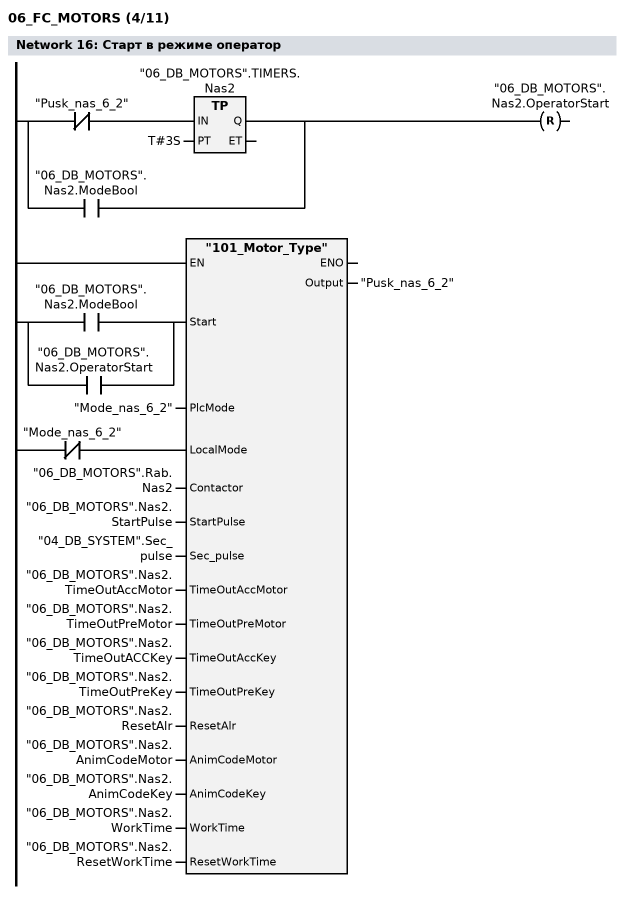
   "06_DB_MOTORS".TIMERS.Nas2.TP(IN := NOT "Pusk_nas_6_2", PT := T#3S);
   IF "06_DB_MOTORS".TIMERS.Nas2.Q OR "06_DB_MOTORS".Nas2.ModeBool THEN
       "06_DB_MOTORS".Nas2.OperatorStart := FALSE;
   END_IF;
   "101_Motor_Type"(Start := "06_DB_MOTORS".Nas2.ModeBool OR "06_DB_MOTORS".Nas2.OperatorStart,
                    PlcMode := "Mode_nas_6_2",
                    LocalMode := NOT "Mode_nas_6_2",
                    Contactor := "06_DB_MOTORS".Rab.Nas2,
                    StartPulse := "06_DB_MOTORS".Nas2.StartPulse,
                    Sec_pulse := "04_DB_SYSTEM".Sec_pulse,
                    TimeOutAccMotor := "06_DB_MOTORS".Nas2.TimeOutAccMotor,
                    TimeOutPreMotor := "06_DB_MOTORS".Nas2.TimeOutPreMotor,
                    TimeOutAccKey := "06_DB_MOTORS".Nas2.TimeOutACCKey,
                    TimeOutPreKey := "06_DB_MOTORS".Nas2.TimeOutPreKey,
                    ResetAlr := "06_DB_MOTORS".Nas2.ResetAlr,
                    AnimCodeMotor := "06_DB_MOTORS".Nas2.AnimCodeMotor,
                    AnimCodeKey := "06_DB_MOTORS".Nas2.AnimCodeKey,
                    WorkTime := "06_DB_MOTORS".Nas2.WorkTime,
                    ResetWorkTime := "06_DB_MOTORS".Nas2.ResetWorkTime,
                    Output => "Pusk_nas_6_2");
END_REGION

REGION Network 17: Старт в режиме оператор
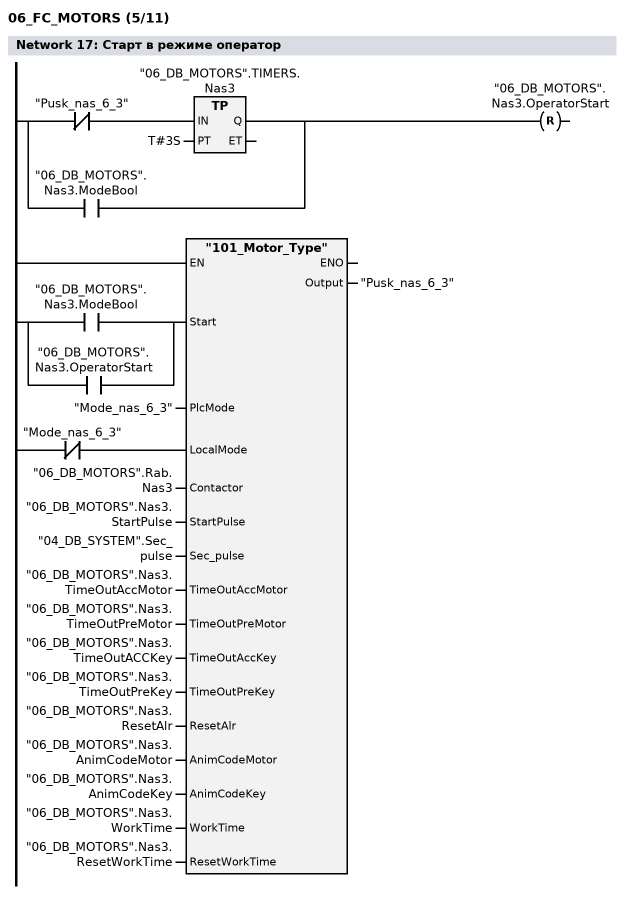
   "06_DB_MOTORS".TIMERS.Nas3.TP(IN := NOT "Pusk_nas_6_3", PT := T#3S);
   IF "06_DB_MOTORS".TIMERS.Nas3.Q OR "06_DB_MOTORS".Nas3.ModeBool THEN
       "06_DB_MOTORS".Nas3.OperatorStart := FALSE;
   END_IF;
   "101_Motor_Type"(Start := "06_DB_MOTORS".Nas3.ModeBool OR "06_DB_MOTORS".Nas3.OperatorStart,
                    PlcMode := "Mode_nas_6_3",
                    LocalMode := NOT "Mode_nas_6_3",
                    Contactor := "06_DB_MOTORS".Rab.Nas3,
                    StartPulse := "06_DB_MOTORS".Nas3.StartPulse,
                    Sec_pulse := "04_DB_SYSTEM".Sec_pulse,
                    TimeOutAccMotor := "06_DB_MOTORS".Nas3.TimeOutAccMotor,
                    TimeOutPreMotor := "06_DB_MOTORS".Nas3.TimeOutPreMotor,
                    TimeOutAccKey := "06_DB_MOTORS".Nas3.TimeOutACCKey,
                    TimeOutPreKey := "06_DB_MOTORS".Nas3.TimeOutPreKey,
                    ResetAlr := "06_DB_MOTORS".Nas3.ResetAlr,
                    AnimCodeMotor := "06_DB_MOTORS".Nas3.AnimCodeMotor,
                    AnimCodeKey := "06_DB_MOTORS".Nas3.AnimCodeKey,
                    WorkTime := "06_DB_MOTORS".Nas3.WorkTime,
                    ResetWorkTime := "06_DB_MOTORS".Nas3.ResetWorkTime,
                    Output => "Pusk_nas_6_3");
END_REGION

REGION Network 18: Старт в режиме оператор
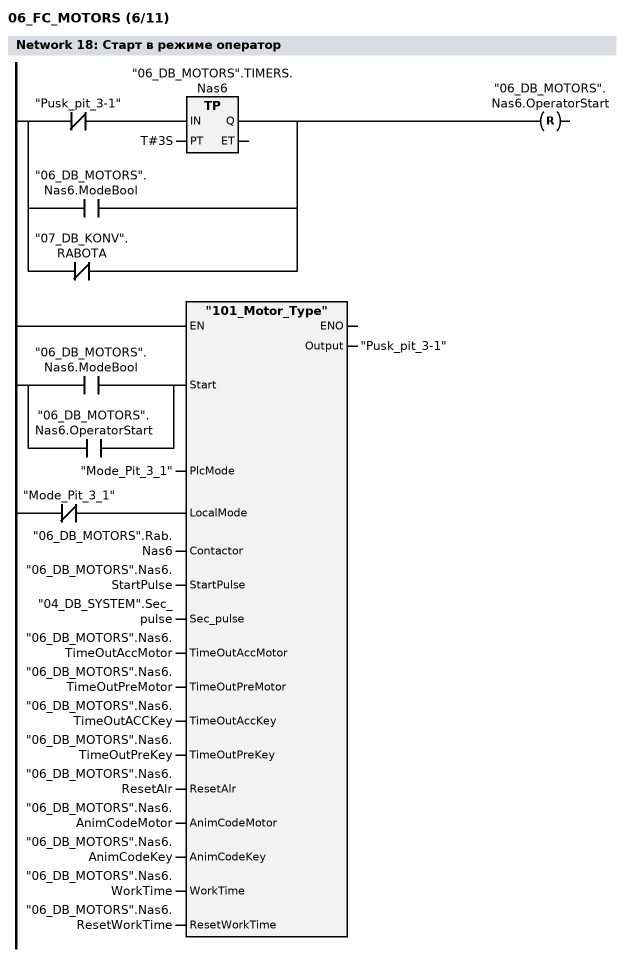
   "06_DB_MOTORS".TIMERS.Nas6.TP(IN := NOT "Pusk_pit_3-1", PT := T#3S);
   IF "06_DB_MOTORS".TIMERS.Nas6.Q OR "06_DB_MOTORS".Nas6.ModeBool OR NOT "07_DB_KONV".RABOTA THEN
       "06_DB_MOTORS".Nas6.OperatorStart := FALSE;
   END_IF;
   "101_Motor_Type"(Start := "06_DB_MOTORS".Nas6.ModeBool OR "06_DB_MOTORS".Nas6.OperatorStart,
                    PlcMode := "Mode_Pit_3_1",
                    LocalMode := NOT "Mode_Pit_3_1",
                    Contactor := "06_DB_MOTORS".Rab.Nas6,
                    StartPulse := "06_DB_MOTORS".Nas6.StartPulse,
                    Sec_pulse := "04_DB_SYSTEM".Sec_pulse,
                    TimeOutAccMotor := "06_DB_MOTORS".Nas6.TimeOutAccMotor,
                    TimeOutPreMotor := "06_DB_MOTORS".Nas6.TimeOutPreMotor,
                    TimeOutAccKey := "06_DB_MOTORS".Nas6.TimeOutACCKey,
                    TimeOutPreKey := "06_DB_MOTORS".Nas6.TimeOutPreKey,
                    ResetAlr := "06_DB_MOTORS".Nas6.ResetAlr,
                    AnimCodeMotor := "06_DB_MOTORS".Nas6.AnimCodeMotor,
                    AnimCodeKey := "06_DB_MOTORS".Nas6.AnimCodeKey,
                    WorkTime := "06_DB_MOTORS".Nas6.WorkTime,
                    ResetWorkTime := "06_DB_MOTORS".Nas6.ResetWorkTime,
                    Output => "Pusk_pit_3-1");
END_REGION

REGION Network 19: Старт в режиме оператор
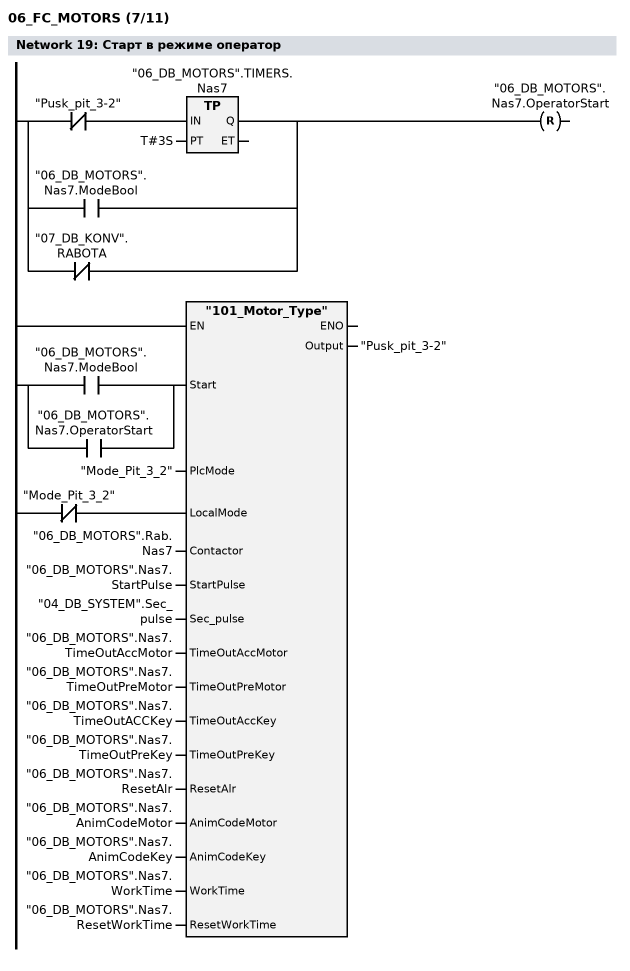
   "06_DB_MOTORS".TIMERS.Nas7.TP(IN := NOT "Pusk_pit_3-2", PT := T#3S);
   IF "06_DB_MOTORS".TIMERS.Nas7.Q OR "06_DB_MOTORS".Nas7.ModeBool OR NOT "07_DB_KONV".RABOTA THEN
       "06_DB_MOTORS".Nas7.OperatorStart := FALSE;
   END_IF;
   "101_Motor_Type"(Start := "06_DB_MOTORS".Nas7.ModeBool OR "06_DB_MOTORS".Nas7.OperatorStart,
                    PlcMode := "Mode_Pit_3_2",
                    LocalMode := NOT "Mode_Pit_3_2",
                    Contactor := "06_DB_MOTORS".Rab.Nas7,
                    StartPulse := "06_DB_MOTORS".Nas7.StartPulse,
                    Sec_pulse := "04_DB_SYSTEM".Sec_pulse,
                    TimeOutAccMotor := "06_DB_MOTORS".Nas7.TimeOutAccMotor,
                    TimeOutPreMotor := "06_DB_MOTORS".Nas7.TimeOutPreMotor,
                    TimeOutAccKey := "06_DB_MOTORS".Nas7.TimeOutACCKey,
                    TimeOutPreKey := "06_DB_MOTORS".Nas7.TimeOutPreKey,
                    ResetAlr := "06_DB_MOTORS".Nas7.ResetAlr,
                    AnimCodeMotor := "06_DB_MOTORS".Nas7.AnimCodeMotor,
                    AnimCodeKey := "06_DB_MOTORS".Nas7.AnimCodeKey,
                    WorkTime := "06_DB_MOTORS".Nas7.WorkTime,
                    ResetWorkTime := "06_DB_MOTORS".Nas7.ResetWorkTime,
                    Output => "Pusk_pit_3-2");
END_REGION

REGION Network 20: Старт в режиме оператор
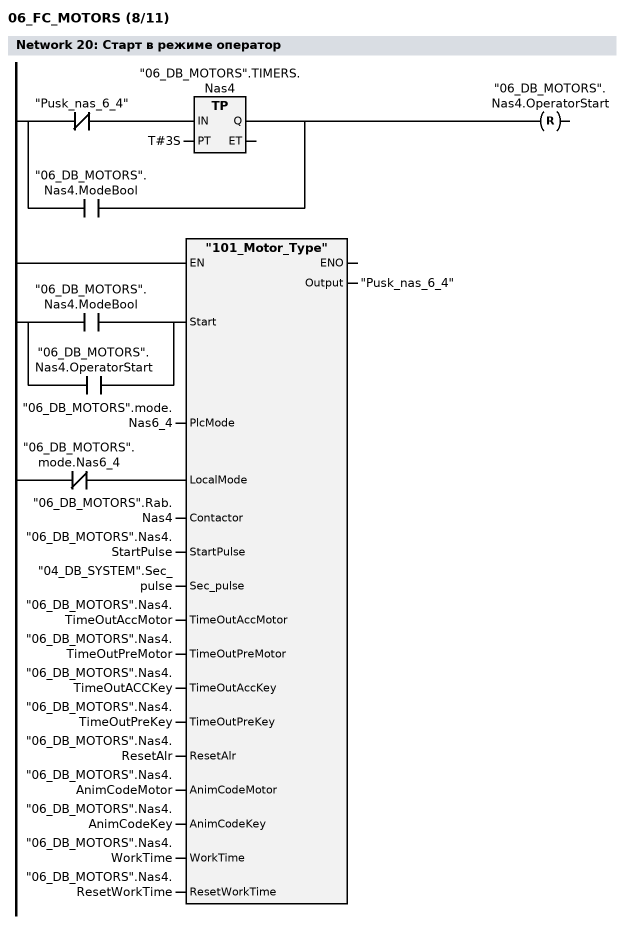
   "06_DB_MOTORS".TIMERS.Nas4.TP(IN := NOT "Pusk_nas_6_4", PT := T#3S);
   IF "06_DB_MOTORS".TIMERS.Nas4.Q OR "06_DB_MOTORS".Nas4.ModeBool THEN
       "06_DB_MOTORS".Nas4.OperatorStart := FALSE;
   END_IF;
   "101_Motor_Type"(Start := "06_DB_MOTORS".Nas4.ModeBool OR "06_DB_MOTORS".Nas4.OperatorStart,
                    PlcMode := "06_DB_MOTORS".mode.Nas6_4,
                    LocalMode := NOT "06_DB_MOTORS".mode.Nas6_4,
                    Contactor := "06_DB_MOTORS".Rab.Nas4,
                    StartPulse := "06_DB_MOTORS".Nas4.StartPulse,
                    Sec_pulse := "04_DB_SYSTEM".Sec_pulse,
                    TimeOutAccMotor := "06_DB_MOTORS".Nas4.TimeOutAccMotor,
                    TimeOutPreMotor := "06_DB_MOTORS".Nas4.TimeOutPreMotor,
                    TimeOutAccKey := "06_DB_MOTORS".Nas4.TimeOutACCKey,
                    TimeOutPreKey := "06_DB_MOTORS".Nas4.TimeOutPreKey,
                    ResetAlr := "06_DB_MOTORS".Nas4.ResetAlr,
                    AnimCodeMotor := "06_DB_MOTORS".Nas4.AnimCodeMotor,
                    AnimCodeKey := "06_DB_MOTORS".Nas4.AnimCodeKey,
                    WorkTime := "06_DB_MOTORS".Nas4.WorkTime,
                    ResetWorkTime := "06_DB_MOTORS".Nas4.ResetWorkTime,
                    Output => "Pusk_nas_6_4");
END_REGION

REGION Network 21: Старт в режиме оператор
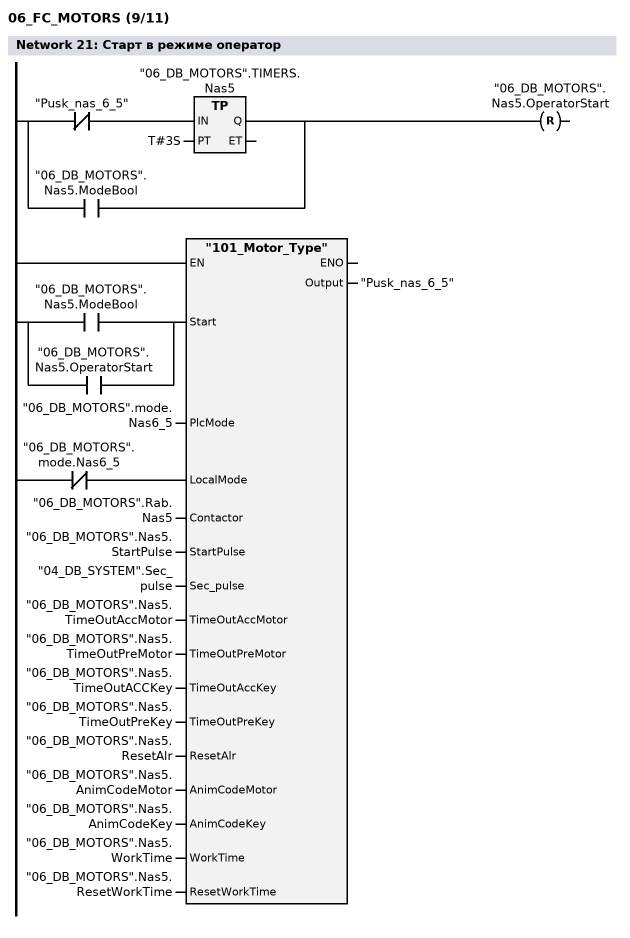
   "06_DB_MOTORS".TIMERS.Nas5.TP(IN := NOT "Pusk_nas_6_5", PT := T#3S);
   IF "06_DB_MOTORS".TIMERS.Nas5.Q OR "06_DB_MOTORS".Nas5.ModeBool THEN
       "06_DB_MOTORS".Nas5.OperatorStart := FALSE;
   END_IF;
   "101_Motor_Type"(Start := "06_DB_MOTORS".Nas5.ModeBool OR "06_DB_MOTORS".Nas5.OperatorStart,
                    PlcMode := "06_DB_MOTORS".mode.Nas6_5,
                    LocalMode := NOT "06_DB_MOTORS".mode.Nas6_5,
                    Contactor := "06_DB_MOTORS".Rab.Nas5,
                    StartPulse := "06_DB_MOTORS".Nas5.StartPulse,
                    Sec_pulse := "04_DB_SYSTEM".Sec_pulse,
                    TimeOutAccMotor := "06_DB_MOTORS".Nas5.TimeOutAccMotor,
                    TimeOutPreMotor := "06_DB_MOTORS".Nas5.TimeOutPreMotor,
                    TimeOutAccKey := "06_DB_MOTORS".Nas5.TimeOutACCKey,
                    TimeOutPreKey := "06_DB_MOTORS".Nas5.TimeOutPreKey,
                    ResetAlr := "06_DB_MOTORS".Nas5.ResetAlr,
                    AnimCodeMotor := "06_DB_MOTORS".Nas5.AnimCodeMotor,
                    AnimCodeKey := "06_DB_MOTORS".Nas5.AnimCodeKey,
                    WorkTime := "06_DB_MOTORS".Nas5.WorkTime,
                    ResetWorkTime := "06_DB_MOTORS".Nas5.ResetWorkTime,
                    Output => "Pusk_nas_6_5");
END_REGION

REGION Network 23: Старт в режиме оператор
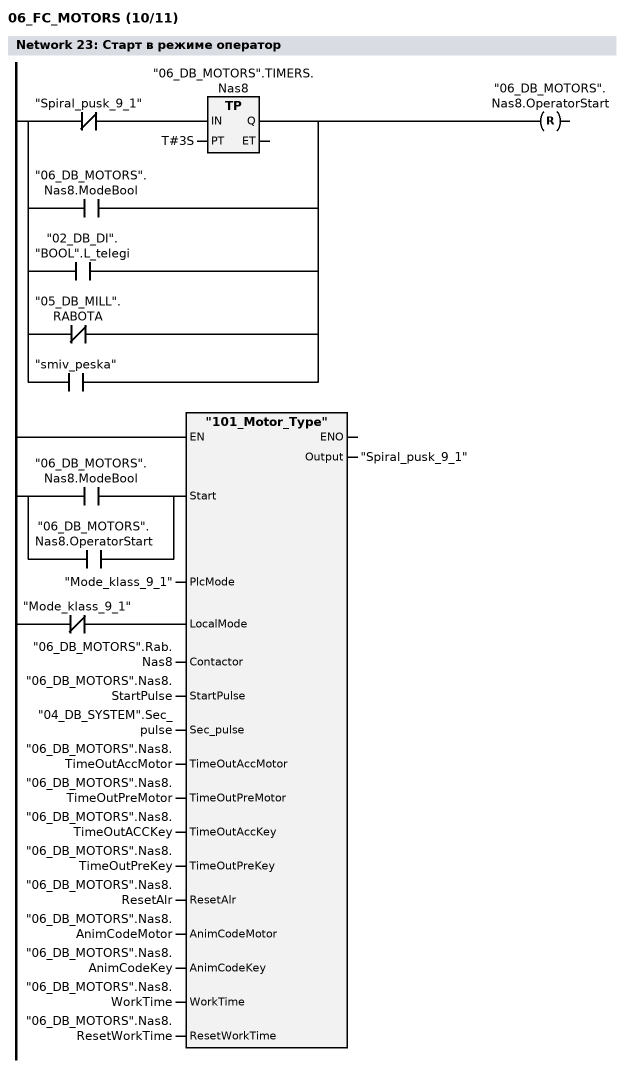
   "06_DB_MOTORS".TIMERS.Nas8.TP(IN := NOT "Spiral_pusk_9_1", PT := T#3S);
   IF "06_DB_MOTORS".TIMERS.Nas8.Q OR "06_DB_MOTORS".Nas8.ModeBool OR "02_DB_DI"."BOOL".L_telegi OR NOT "05_DB_MILL".RABOTA OR "smiv_peska" THEN
       "06_DB_MOTORS".Nas8.OperatorStart := FALSE;
   END_IF;
   "101_Motor_Type"(Start := "06_DB_MOTORS".Nas8.ModeBool OR "06_DB_MOTORS".Nas8.OperatorStart,
                    PlcMode := "Mode_klass_9_1",
                    LocalMode := NOT "Mode_klass_9_1",
                    Contactor := "06_DB_MOTORS".Rab.Nas8,
                    StartPulse := "06_DB_MOTORS".Nas8.StartPulse,
                    Sec_pulse := "04_DB_SYSTEM".Sec_pulse,
                    TimeOutAccMotor := "06_DB_MOTORS".Nas8.TimeOutAccMotor,
                    TimeOutPreMotor := "06_DB_MOTORS".Nas8.TimeOutPreMotor,
                    TimeOutAccKey := "06_DB_MOTORS".Nas8.TimeOutACCKey,
                    TimeOutPreKey := "06_DB_MOTORS".Nas8.TimeOutPreKey,
                    ResetAlr := "06_DB_MOTORS".Nas8.ResetAlr,
                    AnimCodeMotor := "06_DB_MOTORS".Nas8.AnimCodeMotor,
                    AnimCodeKey := "06_DB_MOTORS".Nas8.AnimCodeKey,
                    WorkTime := "06_DB_MOTORS".Nas8.WorkTime,
                    ResetWorkTime := "06_DB_MOTORS".Nas8.ResetWorkTime,
                    Output => "Spiral_pusk_9_1");
END_REGION

REGION Network 24: Старт в режиме оператор
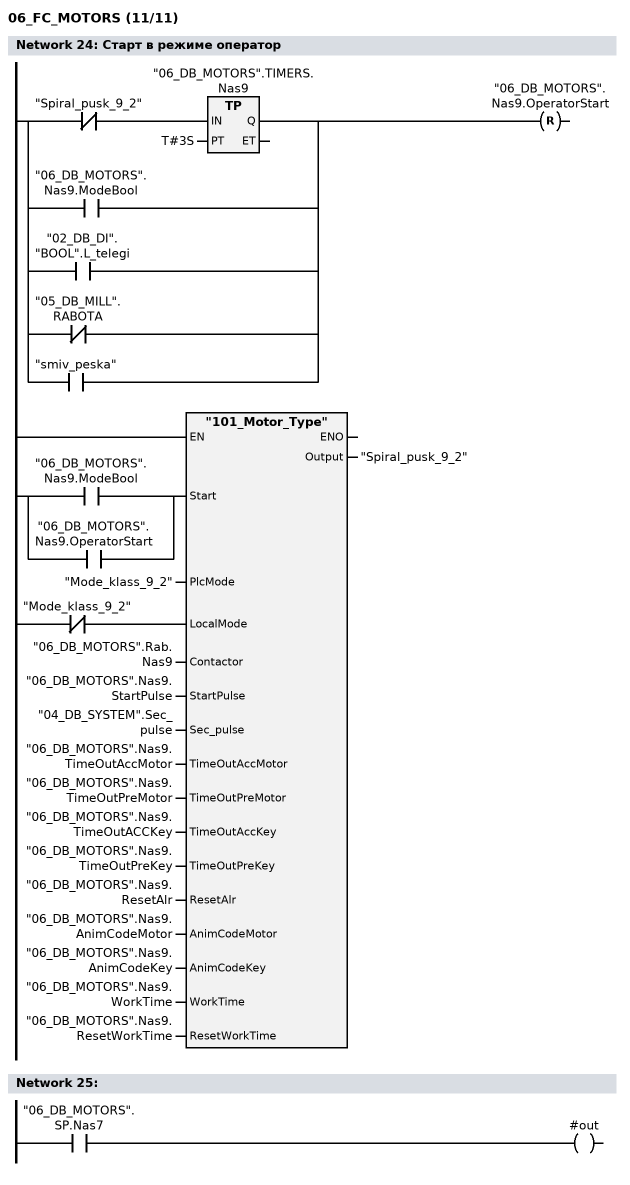
   "06_DB_MOTORS".TIMERS.Nas9.TP(IN := NOT "Spiral_pusk_9_2", PT := T#3S);
   IF "06_DB_MOTORS".TIMERS.Nas9.Q OR "06_DB_MOTORS".Nas9.ModeBool OR "02_DB_DI"."BOOL".L_telegi OR NOT "05_DB_MILL".RABOTA OR "smiv_peska" THEN
       "06_DB_MOTORS".Nas9.OperatorStart := FALSE;
   END_IF;
   "101_Motor_Type"(Start := "06_DB_MOTORS".Nas9.ModeBool OR "06_DB_MOTORS".Nas9.OperatorStart,
                    PlcMode := "Mode_klass_9_2",
                    LocalMode := NOT "Mode_klass_9_2",
                    Contactor := "06_DB_MOTORS".Rab.Nas9,
                    StartPulse := "06_DB_MOTORS".Nas9.StartPulse,
                    Sec_pulse := "04_DB_SYSTEM".Sec_pulse,
                    TimeOutAccMotor := "06_DB_MOTORS".Nas9.TimeOutAccMotor,
                    TimeOutPreMotor := "06_DB_MOTORS".Nas9.TimeOutPreMotor,
                    TimeOutAccKey := "06_DB_MOTORS".Nas9.TimeOutACCKey,
                    TimeOutPreKey := "06_DB_MOTORS".Nas9.TimeOutPreKey,
                    ResetAlr := "06_DB_MOTORS".Nas9.ResetAlr,
                    AnimCodeMotor := "06_DB_MOTORS".Nas9.AnimCodeMotor,
                    AnimCodeKey := "06_DB_MOTORS".Nas9.AnimCodeKey,
                    WorkTime := "06_DB_MOTORS".Nas9.WorkTime,
                    ResetWorkTime := "06_DB_MOTORS".Nas9.ResetWorkTime,
                    Output => "Spiral_pusk_9_2");
END_REGION

REGION Network 25
   RUNG wire#powerrail
      Contact( "06_DB_MOTORS".SP.Nas7 )
      Coil( #out )
   END_RUNG
   // the same network as SCL:
   #out := "06_DB_MOTORS".SP.Nas7;
END_REGION
END_FUNCTION

FUNCTION "09_alarm" : Void   // FC9, LAD
{ S7_Optimized_Access := 'TRUE' }
VERSION : 0.1
   VAR_TEMP   // added for the SCL form of the ladder/FBD networks
      _w1 : Bool;
      _w2 : Bool;
      _w3 : Bool;
      _w4 : Bool;
      _w5 : Bool;
      _w6 : Bool;
      _w7 : Bool;
      _w8 : Bool;
      _w9 : Bool;
      _w10 : Bool;
      _w11 : Bool;
      _w12 : Bool;
      _w13 : Bool;
      _w14 : Bool;
      _w15 : Bool;
      _w16 : Bool;
   END_VAR
BEGIN

REGION Network 1
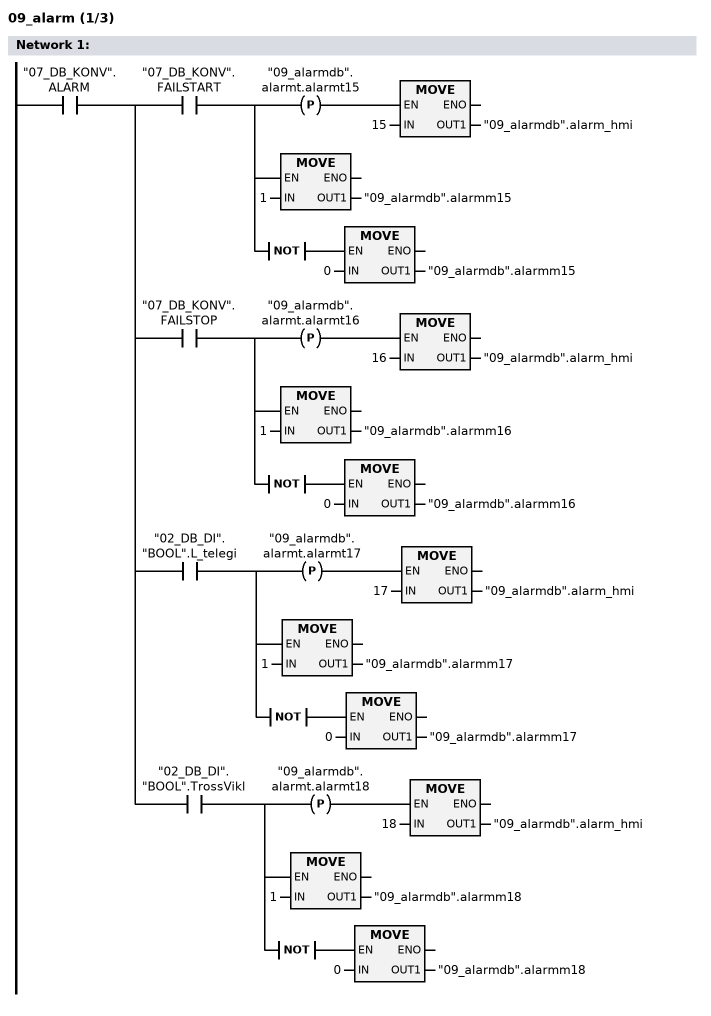
   RUNG wire#powerrail
      Contact( "07_DB_KONV".ALARM )
      wire#w1
      Contact( "07_DB_KONV".FAILSTART )
      wire#w2
      P_Trig( "09_alarmdb".alarmt.alarmt15 )
      Move(in := 15, out1 => "09_alarmdb".alarm_hmi)
   END_RUNG
   RUNG wire#w2
      Move(in := 1, out1 => "09_alarmdb".alarmm15)
   END_RUNG
   RUNG wire#w2
      Not()
      Move(in := 0, out1 => "09_alarmdb".alarmm15)
   END_RUNG
   RUNG wire#w1
      Contact( "07_DB_KONV".FAILSTOP )
      wire#w3
      P_Trig( "09_alarmdb".alarmt.alarmt16 )
      Move(in := 16, out1 => "09_alarmdb".alarm_hmi)
   END_RUNG
   RUNG wire#w3
      Move(in := 1, out1 => "09_alarmdb".alarmm16)
   END_RUNG
   RUNG wire#w3
      Not()
      Move(in := 0, out1 => "09_alarmdb".alarmm16)
   END_RUNG
   RUNG wire#w1
      Contact( "02_DB_DI"."BOOL".L_telegi )
      wire#w4
      P_Trig( "09_alarmdb".alarmt.alarmt17 )
      Move(in := 17, out1 => "09_alarmdb".alarm_hmi)
   END_RUNG
   RUNG wire#w4
      Move(in := 1, out1 => "09_alarmdb".alarmm17)
   END_RUNG
   RUNG wire#w4
      Not()
      Move(in := 0, out1 => "09_alarmdb".alarmm17)
   END_RUNG
   RUNG wire#w1
      Contact( "02_DB_DI"."BOOL".TrossVikl )
      wire#w5
      P_Trig( "09_alarmdb".alarmt.alarmt18 )
      Move(in := 18, out1 => "09_alarmdb".alarm_hmi)
   END_RUNG
   RUNG wire#w5
      Move(in := 1, out1 => "09_alarmdb".alarmm18)
   END_RUNG
   RUNG wire#w5
      Not()
      Move(in := 0, out1 => "09_alarmdb".alarmm18)
   END_RUNG
   // the same network as SCL:
   #_w1 := "07_DB_KONV".ALARM AND "07_DB_KONV".FAILSTART;
   #_w2 := #_w1 AND NOT "09_alarmdb".alarmt.alarmt15;   // rising edge
   "09_alarmdb".alarmt.alarmt15 := #_w1;
   IF #_w2 THEN "09_alarmdb".alarm_hmi := 15; END_IF;
   IF #_w1 THEN "09_alarmdb".alarmm15 := 1; END_IF;
   IF NOT #_w1 THEN "09_alarmdb".alarmm15 := 0; END_IF;
   #_w3 := "07_DB_KONV".ALARM AND "07_DB_KONV".FAILSTOP;
   #_w4 := #_w3 AND NOT "09_alarmdb".alarmt.alarmt16;   // rising edge
   "09_alarmdb".alarmt.alarmt16 := #_w3;
   IF #_w4 THEN "09_alarmdb".alarm_hmi := 16; END_IF;
   IF #_w3 THEN "09_alarmdb".alarmm16 := 1; END_IF;
   IF NOT #_w3 THEN "09_alarmdb".alarmm16 := 0; END_IF;
   #_w5 := "07_DB_KONV".ALARM AND "02_DB_DI"."BOOL".L_telegi;
   #_w6 := #_w5 AND NOT "09_alarmdb".alarmt.alarmt17;   // rising edge
   "09_alarmdb".alarmt.alarmt17 := #_w5;
   IF #_w6 THEN "09_alarmdb".alarm_hmi := 17; END_IF;
   IF #_w5 THEN "09_alarmdb".alarmm17 := 1; END_IF;
   IF NOT #_w5 THEN "09_alarmdb".alarmm17 := 0; END_IF;
   #_w7 := "07_DB_KONV".ALARM AND "02_DB_DI"."BOOL".TrossVikl;
   #_w8 := #_w7 AND NOT "09_alarmdb".alarmt.alarmt18;   // rising edge
   "09_alarmdb".alarmt.alarmt18 := #_w7;
   IF #_w8 THEN "09_alarmdb".alarm_hmi := 18; END_IF;
   IF #_w7 THEN "09_alarmdb".alarmm18 := 1; END_IF;
   IF NOT #_w7 THEN "09_alarmdb".alarmm18 := 0; END_IF;
END_REGION

REGION Network 2
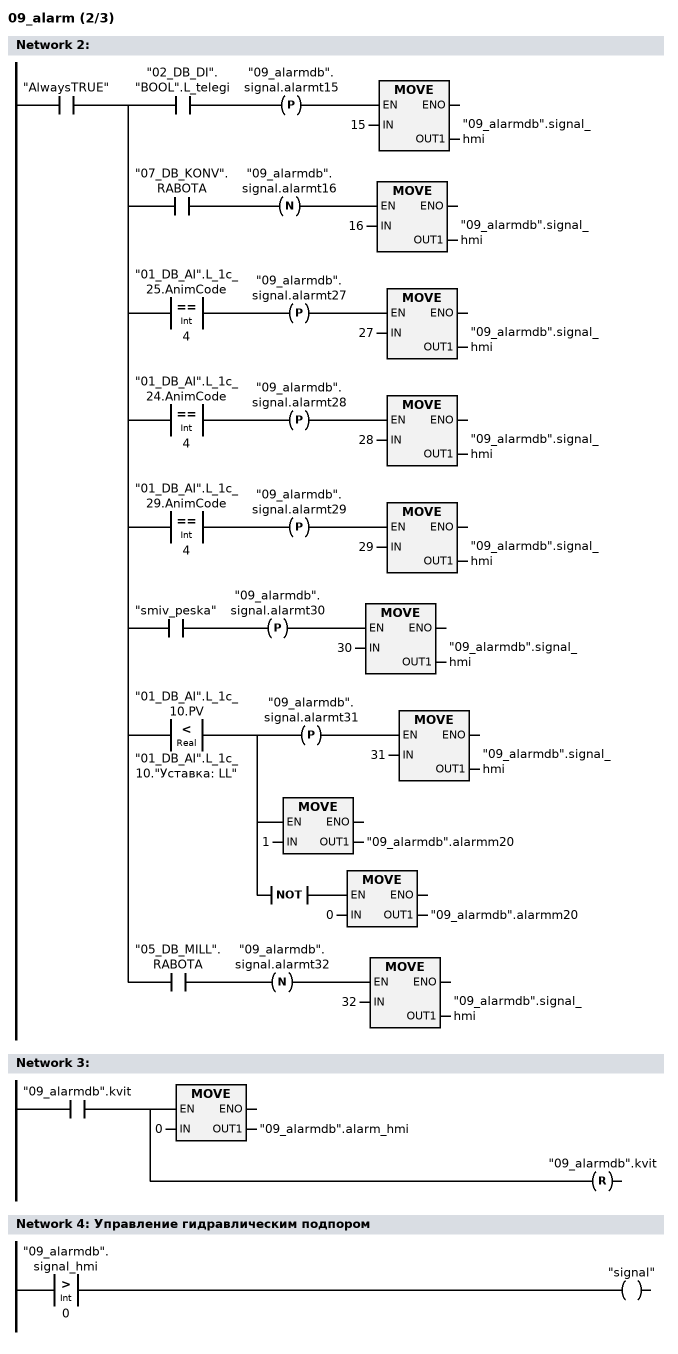
   RUNG wire#powerrail
      Contact( "AlwaysTRUE" )
      wire#w1
      Contact( "02_DB_DI"."BOOL".L_telegi )
      P_Trig( "09_alarmdb".signal.alarmt15 )
      Move(in := 15, out1 => "09_alarmdb".signal_hmi)
   END_RUNG
   RUNG wire#w1
      Contact( "07_DB_KONV".RABOTA )
      N_Trig( "09_alarmdb".signal.alarmt16 )
      Move(in := 16, out1 => "09_alarmdb".signal_hmi)
   END_RUNG
   RUNG wire#w1
      { S7_Templates := "SrcType := Int" } EQ_Contact(in1 := "01_DB_AI".L_1c_25.AnimCode, in2 := 4)
      P_Trig( "09_alarmdb".signal.alarmt27 )
      Move(in := 27, out1 => "09_alarmdb".signal_hmi)
   END_RUNG
   RUNG wire#w1
      { S7_Templates := "SrcType := Int" } EQ_Contact(in1 := "01_DB_AI".L_1c_24.AnimCode, in2 := 4)
      P_Trig( "09_alarmdb".signal.alarmt28 )
      Move(in := 28, out1 => "09_alarmdb".signal_hmi)
   END_RUNG
   RUNG wire#w1
      { S7_Templates := "SrcType := Int" } EQ_Contact(in1 := "01_DB_AI".L_1c_29.AnimCode, in2 := 4)
      P_Trig( "09_alarmdb".signal.alarmt29 )
      Move(in := 29, out1 => "09_alarmdb".signal_hmi)
   END_RUNG
   RUNG wire#w1
      Contact( "smiv_peska" )
      P_Trig( "09_alarmdb".signal.alarmt30 )
      Move(in := 30, out1 => "09_alarmdb".signal_hmi)
   END_RUNG
   RUNG wire#w1
      { S7_Templates := "SrcType := Real" } LT_Contact(in1 := "01_DB_AI".L_1c_10.PV, in2 := "01_DB_AI".L_1c_10."Уставка: LL")
      wire#w2
      P_Trig( "09_alarmdb".signal.alarmt31 )
      Move(in := 31, out1 => "09_alarmdb".signal_hmi)
   END_RUNG
   RUNG wire#w2
      Move(in := 1, out1 => "09_alarmdb".alarmm20)
   END_RUNG
   RUNG wire#w2
      Not()
      Move(in := 0, out1 => "09_alarmdb".alarmm20)
   END_RUNG
   RUNG wire#w1
      Contact( "05_DB_MILL".RABOTA )
      N_Trig( "09_alarmdb".signal.alarmt32 )
      Move(in := 32, out1 => "09_alarmdb".signal_hmi)
   END_RUNG
   // the same network as SCL:
   #_w1 := "AlwaysTRUE" AND "02_DB_DI"."BOOL".L_telegi;
   #_w2 := #_w1 AND NOT "09_alarmdb".signal.alarmt15;   // rising edge
   "09_alarmdb".signal.alarmt15 := #_w1;
   IF #_w2 THEN "09_alarmdb".signal_hmi := 15; END_IF;
   #_w3 := "AlwaysTRUE" AND "07_DB_KONV".RABOTA;
   #_w4 := NOT #_w3 AND "09_alarmdb".signal.alarmt16;   // falling edge
   "09_alarmdb".signal.alarmt16 := #_w3;
   IF #_w4 THEN "09_alarmdb".signal_hmi := 16; END_IF;
   #_w5 := "AlwaysTRUE" AND ("01_DB_AI".L_1c_25.AnimCode = 4);
   #_w6 := #_w5 AND NOT "09_alarmdb".signal.alarmt27;   // rising edge
   "09_alarmdb".signal.alarmt27 := #_w5;
   IF #_w6 THEN "09_alarmdb".signal_hmi := 27; END_IF;
   #_w7 := "AlwaysTRUE" AND ("01_DB_AI".L_1c_24.AnimCode = 4);
   #_w8 := #_w7 AND NOT "09_alarmdb".signal.alarmt28;   // rising edge
   "09_alarmdb".signal.alarmt28 := #_w7;
   IF #_w8 THEN "09_alarmdb".signal_hmi := 28; END_IF;
   #_w9 := "AlwaysTRUE" AND ("01_DB_AI".L_1c_29.AnimCode = 4);
   #_w10 := #_w9 AND NOT "09_alarmdb".signal.alarmt29;   // rising edge
   "09_alarmdb".signal.alarmt29 := #_w9;
   IF #_w10 THEN "09_alarmdb".signal_hmi := 29; END_IF;
   #_w11 := "AlwaysTRUE" AND "smiv_peska";
   #_w12 := #_w11 AND NOT "09_alarmdb".signal.alarmt30;   // rising edge
   "09_alarmdb".signal.alarmt30 := #_w11;
   IF #_w12 THEN "09_alarmdb".signal_hmi := 30; END_IF;
   #_w13 := "AlwaysTRUE" AND ("01_DB_AI".L_1c_10.PV < "01_DB_AI".L_1c_10."Уставка: LL");
   #_w14 := #_w13 AND NOT "09_alarmdb".signal.alarmt31;   // rising edge
   "09_alarmdb".signal.alarmt31 := #_w13;
   IF #_w14 THEN "09_alarmdb".signal_hmi := 31; END_IF;
   IF #_w13 THEN "09_alarmdb".alarmm20 := 1; END_IF;
   IF NOT #_w13 THEN "09_alarmdb".alarmm20 := 0; END_IF;
   #_w15 := "AlwaysTRUE" AND "05_DB_MILL".RABOTA;
   #_w16 := NOT #_w15 AND "09_alarmdb".signal.alarmt32;   // falling edge
   "09_alarmdb".signal.alarmt32 := #_w15;
   IF #_w16 THEN "09_alarmdb".signal_hmi := 32; END_IF;
END_REGION

REGION Network 3
   RUNG wire#powerrail
      Contact( "09_alarmdb".kvit )
      wire#w1
      Move(in := 0, out1 => "09_alarmdb".alarm_hmi)
   END_RUNG
   RUNG wire#w1
      R_Coil( "09_alarmdb".kvit )
   END_RUNG
   // the same network as SCL:
   IF "09_alarmdb".kvit THEN
       "09_alarmdb".alarm_hmi := 0;
       "09_alarmdb".kvit := FALSE;
   END_IF;
END_REGION

REGION Network 4: Управление гидравлическим подпором
   RUNG wire#powerrail
      { S7_Templates := "SrcType := Int" } GT_Contact(in1 := "09_alarmdb".signal_hmi, in2 := 0)
      Coil( "signal" )
   END_RUNG
   // the same network as SCL:
   "signal" := "09_alarmdb".signal_hmi > 0;
END_REGION

REGION Network 5
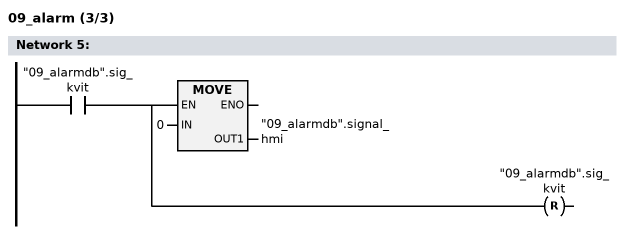
   RUNG wire#powerrail
      Contact( "09_alarmdb".sig_kvit )
      wire#w1
      Move(in := 0, out1 => "09_alarmdb".signal_hmi)
   END_RUNG
   RUNG wire#w1
      R_Coil( "09_alarmdb".sig_kvit )
   END_RUNG
   // the same network as SCL:
   IF "09_alarmdb".sig_kvit THEN
       "09_alarmdb".signal_hmi := 0;
       "09_alarmdb".sig_kvit := FALSE;
   END_IF;
END_REGION
END_FUNCTION

FUNCTION "11_Narabotka" : Void   // FC11, LAD
{ S7_Optimized_Access := 'TRUE' }
VERSION : 0.1
BEGIN

REGION Network 1
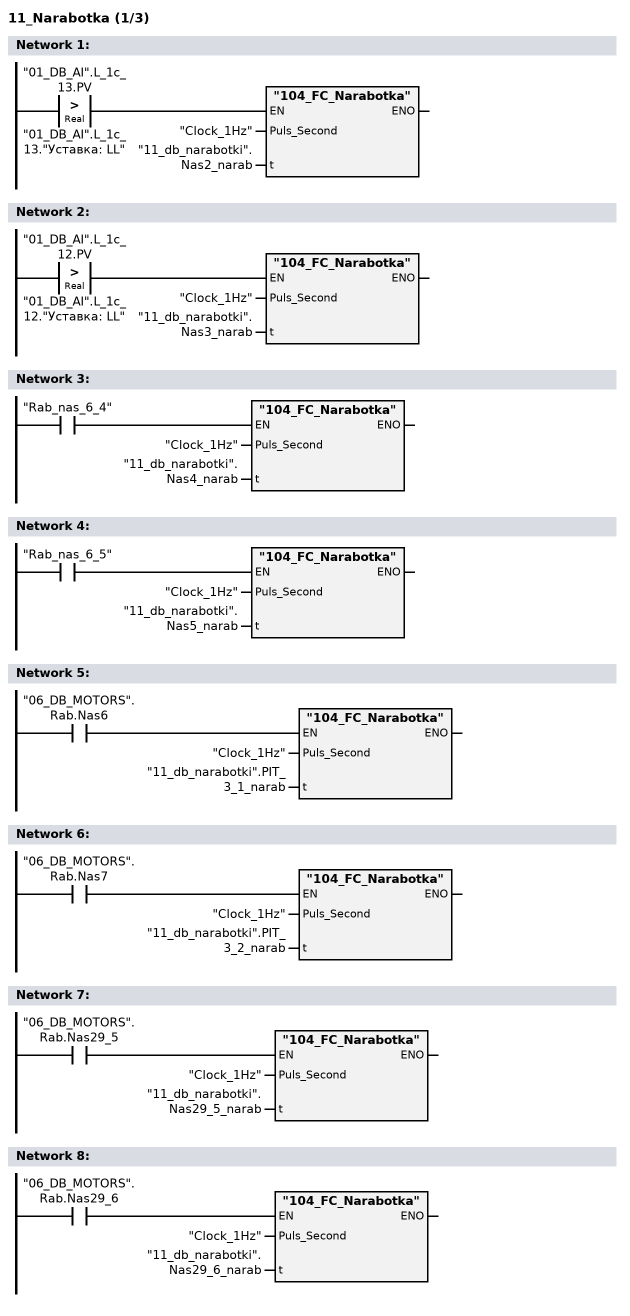
   RUNG wire#powerrail
      { S7_Templates := "SrcType := Real" } GT_Contact(in1 := "01_DB_AI".L_1c_13.PV, in2 := "01_DB_AI".L_1c_13."Уставка: LL")
      "104_FC_Narabotka"(Puls_Second := "Clock_1Hz", t := "11_db_narabotki".Nas2_narab)
   END_RUNG
   // the same network as SCL:
   IF "01_DB_AI".L_1c_13.PV > "01_DB_AI".L_1c_13."Уставка: LL" THEN
       "104_FC_Narabotka"(Puls_Second := "Clock_1Hz", t := "11_db_narabotki".Nas2_narab);
   END_IF;
END_REGION

REGION Network 2
   RUNG wire#powerrail
      { S7_Templates := "SrcType := Real" } GT_Contact(in1 := "01_DB_AI".L_1c_12.PV, in2 := "01_DB_AI".L_1c_12."Уставка: LL")
      "104_FC_Narabotka"(Puls_Second := "Clock_1Hz", t := "11_db_narabotki".Nas3_narab)
   END_RUNG
   // the same network as SCL:
   IF "01_DB_AI".L_1c_12.PV > "01_DB_AI".L_1c_12."Уставка: LL" THEN
       "104_FC_Narabotka"(Puls_Second := "Clock_1Hz", t := "11_db_narabotki".Nas3_narab);
   END_IF;
END_REGION

REGION Network 3
   RUNG wire#powerrail
      Contact( "Rab_nas_6_4" )
      "104_FC_Narabotka"(Puls_Second := "Clock_1Hz", t := "11_db_narabotki".Nas4_narab)
   END_RUNG
   // the same network as SCL:
   IF "Rab_nas_6_4" THEN
       "104_FC_Narabotka"(Puls_Second := "Clock_1Hz", t := "11_db_narabotki".Nas4_narab);
   END_IF;
END_REGION

REGION Network 4
   RUNG wire#powerrail
      Contact( "Rab_nas_6_5" )
      "104_FC_Narabotka"(Puls_Second := "Clock_1Hz", t := "11_db_narabotki".Nas5_narab)
   END_RUNG
   // the same network as SCL:
   IF "Rab_nas_6_5" THEN
       "104_FC_Narabotka"(Puls_Second := "Clock_1Hz", t := "11_db_narabotki".Nas5_narab);
   END_IF;
END_REGION

REGION Network 5
   RUNG wire#powerrail
      Contact( "06_DB_MOTORS".Rab.Nas6 )
      "104_FC_Narabotka"(Puls_Second := "Clock_1Hz", t := "11_db_narabotki".PIT_3_1_narab)
   END_RUNG
   // the same network as SCL:
   IF "06_DB_MOTORS".Rab.Nas6 THEN
       "104_FC_Narabotka"(Puls_Second := "Clock_1Hz", t := "11_db_narabotki".PIT_3_1_narab);
   END_IF;
END_REGION

REGION Network 6
   RUNG wire#powerrail
      Contact( "06_DB_MOTORS".Rab.Nas7 )
      "104_FC_Narabotka"(Puls_Second := "Clock_1Hz", t := "11_db_narabotki".PIT_3_2_narab)
   END_RUNG
   // the same network as SCL:
   IF "06_DB_MOTORS".Rab.Nas7 THEN
       "104_FC_Narabotka"(Puls_Second := "Clock_1Hz", t := "11_db_narabotki".PIT_3_2_narab);
   END_IF;
END_REGION

REGION Network 7
   RUNG wire#powerrail
      Contact( "06_DB_MOTORS".Rab.Nas29_5 )
      "104_FC_Narabotka"(Puls_Second := "Clock_1Hz", t := "11_db_narabotki".Nas29_5_narab)
   END_RUNG
   // the same network as SCL:
   IF "06_DB_MOTORS".Rab.Nas29_5 THEN
       "104_FC_Narabotka"(Puls_Second := "Clock_1Hz", t := "11_db_narabotki".Nas29_5_narab);
   END_IF;
END_REGION

REGION Network 8
   RUNG wire#powerrail
      Contact( "06_DB_MOTORS".Rab.Nas29_6 )
      "104_FC_Narabotka"(Puls_Second := "Clock_1Hz", t := "11_db_narabotki".Nas29_6_narab)
   END_RUNG
   // the same network as SCL:
   IF "06_DB_MOTORS".Rab.Nas29_6 THEN
       "104_FC_Narabotka"(Puls_Second := "Clock_1Hz", t := "11_db_narabotki".Nas29_6_narab);
   END_IF;
END_REGION

REGION Network 9
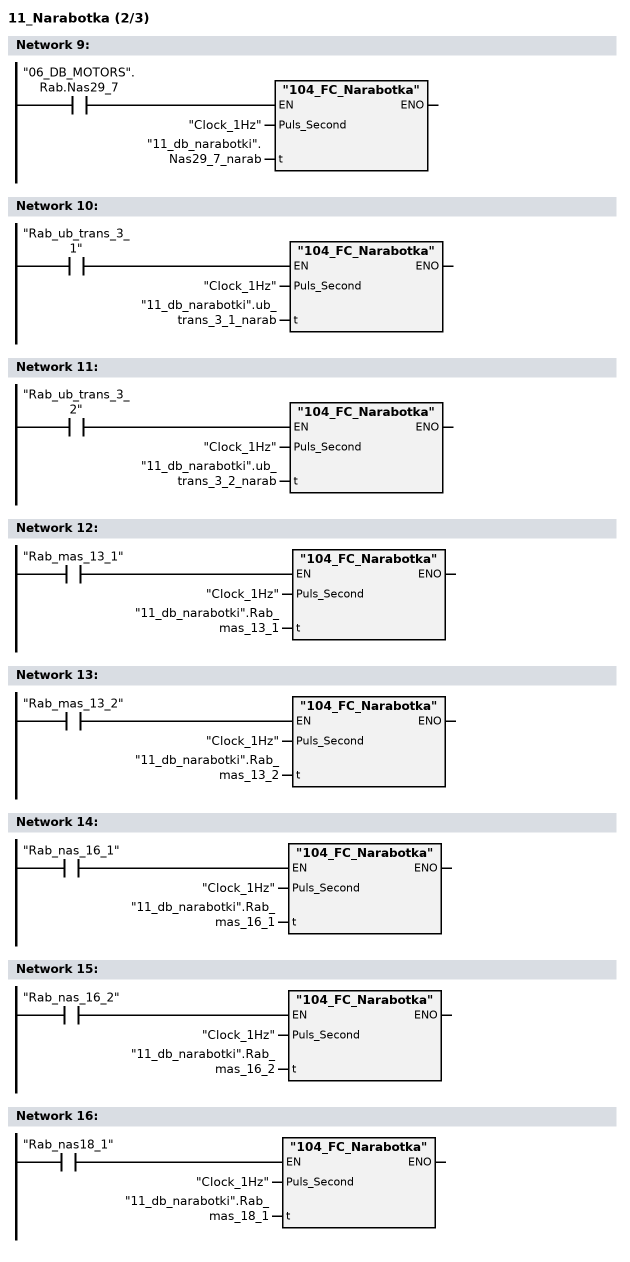
   RUNG wire#powerrail
      Contact( "06_DB_MOTORS".Rab.Nas29_7 )
      "104_FC_Narabotka"(Puls_Second := "Clock_1Hz", t := "11_db_narabotki".Nas29_7_narab)
   END_RUNG
   // the same network as SCL:
   IF "06_DB_MOTORS".Rab.Nas29_7 THEN
       "104_FC_Narabotka"(Puls_Second := "Clock_1Hz", t := "11_db_narabotki".Nas29_7_narab);
   END_IF;
END_REGION

REGION Network 10
   RUNG wire#powerrail
      Contact( "Rab_ub_trans_3_1" )
      "104_FC_Narabotka"(Puls_Second := "Clock_1Hz", t := "11_db_narabotki".ub_trans_3_1_narab)
   END_RUNG
   // the same network as SCL:
   IF "Rab_ub_trans_3_1" THEN
       "104_FC_Narabotka"(Puls_Second := "Clock_1Hz", t := "11_db_narabotki".ub_trans_3_1_narab);
   END_IF;
END_REGION

REGION Network 11
   RUNG wire#powerrail
      Contact( "Rab_ub_trans_3_2" )
      "104_FC_Narabotka"(Puls_Second := "Clock_1Hz", t := "11_db_narabotki".ub_trans_3_2_narab)
   END_RUNG
   // the same network as SCL:
   IF "Rab_ub_trans_3_2" THEN
       "104_FC_Narabotka"(Puls_Second := "Clock_1Hz", t := "11_db_narabotki".ub_trans_3_2_narab);
   END_IF;
END_REGION

REGION Network 12
   RUNG wire#powerrail
      Contact( "Rab_mas_13_1" )
      "104_FC_Narabotka"(Puls_Second := "Clock_1Hz", t := "11_db_narabotki".Rab_mas_13_1)
   END_RUNG
   // the same network as SCL:
   IF "Rab_mas_13_1" THEN
       "104_FC_Narabotka"(Puls_Second := "Clock_1Hz", t := "11_db_narabotki".Rab_mas_13_1);
   END_IF;
END_REGION

REGION Network 13
   RUNG wire#powerrail
      Contact( "Rab_mas_13_2" )
      "104_FC_Narabotka"(Puls_Second := "Clock_1Hz", t := "11_db_narabotki".Rab_mas_13_2)
   END_RUNG
   // the same network as SCL:
   IF "Rab_mas_13_2" THEN
       "104_FC_Narabotka"(Puls_Second := "Clock_1Hz", t := "11_db_narabotki".Rab_mas_13_2);
   END_IF;
END_REGION

REGION Network 14
   RUNG wire#powerrail
      Contact( "Rab_nas_16_1" )
      "104_FC_Narabotka"(Puls_Second := "Clock_1Hz", t := "11_db_narabotki".Rab_mas_16_1)
   END_RUNG
   // the same network as SCL:
   IF "Rab_nas_16_1" THEN
       "104_FC_Narabotka"(Puls_Second := "Clock_1Hz", t := "11_db_narabotki".Rab_mas_16_1);
   END_IF;
END_REGION

REGION Network 15
   RUNG wire#powerrail
      Contact( "Rab_nas_16_2" )
      "104_FC_Narabotka"(Puls_Second := "Clock_1Hz", t := "11_db_narabotki".Rab_mas_16_2)
   END_RUNG
   // the same network as SCL:
   IF "Rab_nas_16_2" THEN
       "104_FC_Narabotka"(Puls_Second := "Clock_1Hz", t := "11_db_narabotki".Rab_mas_16_2);
   END_IF;
END_REGION

REGION Network 16
   RUNG wire#powerrail
      Contact( "Rab_nas18_1" )
      "104_FC_Narabotka"(Puls_Second := "Clock_1Hz", t := "11_db_narabotki".Rab_mas_18_1)
   END_RUNG
   // the same network as SCL:
   IF "Rab_nas18_1" THEN
       "104_FC_Narabotka"(Puls_Second := "Clock_1Hz", t := "11_db_narabotki".Rab_mas_18_1);
   END_IF;
END_REGION

REGION Network 17
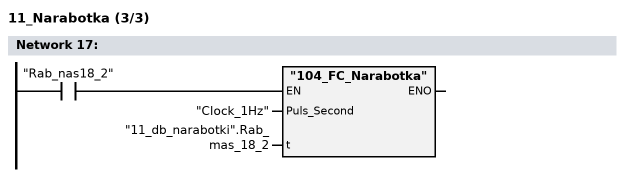
   RUNG wire#powerrail
      Contact( "Rab_nas18_2" )
      "104_FC_Narabotka"(Puls_Second := "Clock_1Hz", t := "11_db_narabotki".Rab_mas_18_2)
   END_RUNG
   // the same network as SCL:
   IF "Rab_nas18_2" THEN
       "104_FC_Narabotka"(Puls_Second := "Clock_1Hz", t := "11_db_narabotki".Rab_mas_18_2);
   END_IF;
END_REGION
END_FUNCTION

FUNCTION "100_Analog_Type" : Void   // FC100, LAD
TITLE = Блок обработки сигнала аналогового входа 4-20мА
{ S7_Optimized_Access := 'FALSE' }
VERSION : 0.1
   VAR_INPUT
      Вход : Int;
   END_VAR
   VAR_IN_OUT
      HMI : "AI_STR";
   END_VAR
   VAR_TEMP
      Val_temp : Real;
   END_VAR
   VAR CONSTANT
      Undershoot_MIN : Int := -4864;   // Минимальная граница Недолёт
      Overshoot_MAX : Int := 32511;   // Минимальная граница Перелет
      Underflow : Int := -32768;   // Обрыв
      Overflow : Int := 32767;   // Зашкал
   END_VAR
BEGIN

REGION Network 1: Вычисление тока в мА
